(* Logix 5000 project; controller PLC_MCC1300_75F1 vendor 1 type 14 code 166 rev 32.11; software revision 32.04; part 74 of 83 *)
(* tags used below, declared in another part *)
   AUX_tConvoyCap_ZC_NULL : UDT_ConvoyCap_ZC;
   CONST_rgdDestMask : DINT[32];   // Destination Mask
   CONST_tAux : AUX_COSTANTS;
   CONST_tPlant : UDT_PLANT_CONSTANTS;
   GP_PosWindow : GP_PosWindow;
   GP_TrackingAddCap : GP_TrackingAddCap;
   M302SpeedUp : MAC_SpeedUp;
   M303_dHalfWidthDifference : DINT;
   M307ASpeedUp : MAC_SpeedUp;
   M30xTrimDeck : MAC_TrimmingDeck[5];
   M30xTrimDeck_DATA : UDT_ConvoyCap_ZC[5];
   M30xTrimDeck_HMR : MAC_TrimmingDeck_HMR[5];
   M30xTrimDeck_HMW : MAC_TrimmingDeck_HMW[5];
   M30xTrimWheel : MAC_TrimmingWheels[5];
   M310Popup : MAC_Popup_ZC[2];
   M315Popup : MAC_Popup_ZC[2];
   M350Popup : MAC_Popup_ZC;
   O : INT[128];
   Sbr_IN_dCapIndex : DINT;
   Sbr_IN_DestinationCullet : DINT;
   Sbr_IN_dIndexHead : DINT;
   Sbr_IN_ReentryPosition : DINT;
   Sbr_IN_ReentryPosition_max : DINT;
   Sbr_IN_ReentryPosition_min : DINT;
   Sbr_INO_DestinationLite : DINT;
   Sbr_INO_tConvoy_SL : UDT_Convoy_SL;
   Sbr_INO_tConvoyCap_ZC : UDT_ConvoyCap_ZC;
   Sbr_INO_xALLForDestination : BOOL;
   Sbr_INO_xAllLiteToCullet : BOOL;
   Sbr_INO_xAtLeastOneForDestination : BOOL;
   Sbr_INO_xAtLeastOneToCullet : BOOL;
   Sbr_OUT_dTotalCaps : DINT;
   Sbr_OUT_rgdConvoyGaps : DINT[4];
   Sbr_OUT_rgdConvoyLengths : DINT[4];
   TMP_d : DINT;
   TMP_dCap : DINT;
   TMP_dConvoySearchMax : DINT;
   TMP_dIndC : DINT;
   TMP_dIndex : DINT;
   TMP_dLite : DINT;
   TMP_dManualTargetPos : DINT;
   TMP_dMaxCap : DINT;
   TMP_dMaxLite : DINT;
   TMP_dNextCap : DINT;
   TMP_dPointer : DINT;
   TMP_dWander : DINT;
   TMP_rgdIndexC : DINT[4];
   TMP_rgdPnt : DINT[5];
   TMP_x : BOOL;
   TMP_xDebugOFF : BOOL;
   TMP_xDebugON : BOOL;
   xAlwaysOFF : BOOL;
   xAlwaysON : BOOL;
   Z200_SnapDataEth : UDT_ConvoyCap_ZC[2];
   Z300_BufferPlate : UDT_LINE_BUFFER_PLATE;
   Z300_Conveyor_Conf : UDT_Conveyor_Config[29];
   Z300_dEndTrackingPosition : DINT;
   Z300_LineTracking : UDT_LINE_TRACKING;
   Z301 : MAC_Zone_ML;
   Z401_HMI_rgtPlateScada : HMI_LiteData[5,2,7];
   Z401_HMI_rgtPlateScada_Internal : HMI_LiteData[5,2,7];
   Z402_HMI_rgtPlateScada : HMI_LiteData[5,2,7];
   Z402_HMI_rgtPlateScada_Internal : HMI_LiteData[5,2,7];
   Z900_HMI_rgtPlateScada : HMI_LiteData[5,2,7];
   Z900_HMI_rgtPlateScada_Internal : HMI_LiteData[5,2,7];
(* MainProgram, continued *)

ROUTINE Machines_Config   (* structured text *)
   //// MACHINES CONFIGURATION ////
   
   //M302 Speed-Up
   M302SpeedUp.AUX_dConveyorLength_cmm := 0;
   FOR TMP_dIndex := 0 TO 9 DO
   	M302SpeedUp.AUX_dConveyorLength_cmm := M302SpeedUp.AUX_dConveyorLength_cmm + Z300_Conveyor_Conf[TMP_dIndex].dLengthConveyor_cmm;
   END_FOR;
   
   //M302 Trim Deck
   M30xTrimDeck[0].CONF_dAutoSpeed_mm_min := 1000; //1680 //1000 (/60)
   M30xTrimDeck[0].CONF_dManualSpeed_mm_min := 300; //500 //900 //300 (/60)
   M30xTrimDeck[0].CONF_dConveyorLength_cmm := Z300_LineTracking.rgtTrkConv[2].dLengthConveyor + Z300_LineTracking.rgtTrkConv[3].dLengthConveyor + Z300_LineTracking.rgtTrkConv[4].dLengthConveyor + Z300_LineTracking.rgtTrkConv[5].dLengthConveyor + Z300_LineTracking.rgtTrkConv[6].dLengthConveyor;
   M30xTrimDeck[0].CONF_dStartPositionFrame := Z300_LineTracking.rgtTrkConv[2].dStartPosition_cmm;
   M30xTrimDeck[0].CONF_dStopPositionFrame_cmm := Z300_LineTracking.rgtTrkConv[6].dEndPosition_cmm;
   M30xTrimDeck[0].CONF_dTrimDeckPreset[0] := 2055; //mm
   M30xTrimDeck[0].CONF_dTrimDeckPreset[1] := 2055; //mm
   M30xTrimDeck[0].CONF_dTrimDeckCleanPos_cmm[0] := 205500;
   M30xTrimDeck[0].CONF_dTrimDeckCleanPos_cmm[1] := 205500;
   M30xTrimDeck[0].CONF_dMaxTimeToReachPosition_ms := 600;
   M30xTrimDeck[0].CONF_dTolerance_cmm := 200;
   M30xTrimDeck[0].CONF_dTrimDeckTargetWindow_cmm[0] := 200;
   M30xTrimDeck[0].CONF_dTrimDeckTargetWindow_cmm[1] := 200;
   M30xTrimDeck[0].CONF_rAcceleration_m_s2[0] := 0.06;
   M30xTrimDeck[0].CONF_rDeceleration_m_s2[0] := 0.06;
   M30xTrimDeck[0].CONF_rAcceleration_m_s2[1] := 0.06;
   M30xTrimDeck[0].CONF_rDeceleration_m_s2[1] := 0.06;
   M30xTrimDeck[0].tmOF_DriveEnable[0].PRE := 30000;
   M30xTrimDeck[0].tmOF_DriveEnable[1].PRE := 30000;
   M30xTrimDeck[0].tmON_FeedbackTimeOut[0].PRE := 5000;
   M30xTrimDeck[0].tmON_FeedbackTimeOut[1].PRE := 5000;
   M30xTrimDeck[0].tmON_FeedbackDriveReady[0].PRE := 1000;
   M30xTrimDeck[0].tmON_FeedbackDriveReady[1].PRE := 1000;
   
   //M303 Trim Deck
   M30xTrimDeck[1].CONF_dAutoSpeed_mm_min := 1000; //1680 //1000 (/60)
   M30xTrimDeck[1].CONF_dManualSpeed_mm_min := 300; //500 //900 //300 (/60)
   M30xTrimDeck[1].CONF_dConveyorLength_cmm := Z300_LineTracking.rgtTrkConv[7].dLengthConveyor + Z300_LineTracking.rgtTrkConv[8].dLengthConveyor;
   M30xTrimDeck[1].CONF_dStartPositionFrame := Z300_LineTracking.rgtTrkConv[7].dStartPosition_cmm;
   M30xTrimDeck[1].CONF_dStopPositionFrame_cmm := Z300_LineTracking.rgtTrkConv[8].dEndPosition_cmm;
   M30xTrimDeck[1].CONF_dTrimDeckPreset[0] := 2055; //mm
   M30xTrimDeck[1].CONF_dTrimDeckPreset[1] := 2055; //mm
   M30xTrimDeck[1].CONF_dTrimDeckCleanPos_cmm[0] := 205500;
   M30xTrimDeck[1].CONF_dTrimDeckCleanPos_cmm[1] := 205500;
   M30xTrimDeck[1].CONF_dMaxTimeToReachPosition_ms := 600;
   M30xTrimDeck[1].CONF_dTolerance_cmm := 200;
   M30xTrimDeck[1].CONF_dTrimDeckTargetWindow_cmm[0] := 200;
   M30xTrimDeck[1].CONF_dTrimDeckTargetWindow_cmm[1] := 200;
   M30xTrimDeck[1].CONF_rAcceleration_m_s2[0] := 0.06;
   M30xTrimDeck[1].CONF_rDeceleration_m_s2[0] := 0.06;
   M30xTrimDeck[1].CONF_rAcceleration_m_s2[1] := 0.06;
   M30xTrimDeck[1].CONF_rDeceleration_m_s2[1] := 0.06;
   M30xTrimDeck[1].tmOF_DriveEnable[0].PRE := 30000;
   M30xTrimDeck[1].tmOF_DriveEnable[1].PRE := 30000;
   M30xTrimDeck[1].tmON_FeedbackTimeOut[0].PRE := 5000;
   M30xTrimDeck[1].tmON_FeedbackTimeOut[1].PRE := 5000;
   M30xTrimDeck[1].tmON_FeedbackDriveReady[0].PRE := 1000;
   M30xTrimDeck[1].tmON_FeedbackDriveReady[1].PRE := 1000;
   
   //M304 Trim Deck
   M30xTrimDeck[2].CONF_dAutoSpeed_mm_min := 1000; //1680 //1000 (/60)
   M30xTrimDeck[2].CONF_dManualSpeed_mm_min := 300; //500 //900 //300 (/60)
   M30xTrimDeck[2].CONF_dConveyorLength_cmm := Z300_LineTracking.rgtTrkConv[9].dLengthConveyor;
   M30xTrimDeck[2].CONF_dStartPositionFrame := Z300_LineTracking.rgtTrkConv[9].dStartPosition_cmm;
   M30xTrimDeck[2].CONF_dStopPositionFrame_cmm := Z300_LineTracking.rgtTrkConv[9].dEndPosition_cmm;
   M30xTrimDeck[2].CONF_dTrimDeckPreset[0] := 2055; //mm
   M30xTrimDeck[2].CONF_dTrimDeckPreset[1] := 2055; //mm
   M30xTrimDeck[2].CONF_dTrimDeckCleanPos_cmm[0] := 205500;
   M30xTrimDeck[2].CONF_dTrimDeckCleanPos_cmm[1] := 205500;
   M30xTrimDeck[2].CONF_dMaxTimeToReachPosition_ms := 600;
   M30xTrimDeck[2].CONF_dTolerance_cmm := 200;
   M30xTrimDeck[2].CONF_dTrimDeckTargetWindow_cmm[0] := 200;
   M30xTrimDeck[2].CONF_dTrimDeckTargetWindow_cmm[1] := 200;
   M30xTrimDeck[2].CONF_rAcceleration_m_s2[0] := 0.06;
   M30xTrimDeck[2].CONF_rDeceleration_m_s2[0] := 0.06;
   M30xTrimDeck[2].CONF_rAcceleration_m_s2[1] := 0.06;
   M30xTrimDeck[2].CONF_rDeceleration_m_s2[1] := 0.06;
   M30xTrimDeck[2].tmOF_DriveEnable[0].PRE := 30000;
   M30xTrimDeck[2].tmOF_DriveEnable[1].PRE := 30000;
   M30xTrimDeck[2].tmON_FeedbackTimeOut[0].PRE := 5000;
   M30xTrimDeck[2].tmON_FeedbackTimeOut[1].PRE := 5000;
   M30xTrimDeck[2].tmON_FeedbackDriveReady[0].PRE := 1000;
   M30xTrimDeck[2].tmON_FeedbackDriveReady[1].PRE := 1000;
   
   //M305 Trim Deck
   M30xTrimDeck[3].CONF_dAutoSpeed_mm_min := 1000; //1680 //1000 (/60)
   M30xTrimDeck[3].CONF_dManualSpeed_mm_min := 300; //500 //900 //300 (/60)
   M30xTrimDeck[3].CONF_dConveyorLength_cmm := Z300_LineTracking.rgtTrkConv[10].dLengthConveyor;
   M30xTrimDeck[3].CONF_dStartPositionFrame := Z300_LineTracking.rgtTrkConv[10].dStartPosition_cmm;
   M30xTrimDeck[3].CONF_dStopPositionFrame_cmm := Z300_LineTracking.rgtTrkConv[10].dEndPosition_cmm;
   M30xTrimDeck[3].CONF_dTrimDeckPreset[0] := 2055; //mm
   M30xTrimDeck[3].CONF_dTrimDeckPreset[1] := 2055; //mm
   M30xTrimDeck[3].CONF_dTrimDeckCleanPos_cmm[0] := 205500;
   M30xTrimDeck[3].CONF_dTrimDeckCleanPos_cmm[1] := 205500;
   M30xTrimDeck[3].CONF_dMaxTimeToReachPosition_ms := 600;
   M30xTrimDeck[3].CONF_dTolerance_cmm := 200;
   M30xTrimDeck[3].CONF_dTrimDeckTargetWindow_cmm[0] := 200;
   M30xTrimDeck[3].CONF_dTrimDeckTargetWindow_cmm[1] := 200;
   M30xTrimDeck[3].CONF_rAcceleration_m_s2[0] := 0.06;
   M30xTrimDeck[3].CONF_rDeceleration_m_s2[0] := 0.06;
   M30xTrimDeck[3].CONF_rAcceleration_m_s2[1] := 0.06;
   M30xTrimDeck[3].CONF_rDeceleration_m_s2[1] := 0.06;
   M30xTrimDeck[3].tmOF_DriveEnable[0].PRE := 30000;
   M30xTrimDeck[3].tmOF_DriveEnable[1].PRE := 30000;
   M30xTrimDeck[3].tmON_FeedbackTimeOut[0].PRE := 5000;
   M30xTrimDeck[3].tmON_FeedbackTimeOut[1].PRE := 5000;
   M30xTrimDeck[3].tmON_FeedbackDriveReady[0].PRE := 1000;
   M30xTrimDeck[3].tmON_FeedbackDriveReady[1].PRE := 1000;
   
   //M306 Trim Deck
   M30xTrimDeck[4].CONF_dAutoSpeed_mm_min := 1000; //1680 //1000 (/60)
   M30xTrimDeck[4].CONF_dManualSpeed_mm_min := 300; //500 //900 //300 (/60)
   M30xTrimDeck[4].CONF_dConveyorLength_cmm := Z300_LineTracking.rgtTrkConv[11].dLengthConveyor;
   M30xTrimDeck[4].CONF_dStartPositionFrame := Z300_LineTracking.rgtTrkConv[11].dStartPosition_cmm;
   M30xTrimDeck[4].CONF_dStopPositionFrame_cmm := Z300_LineTracking.rgtTrkConv[11].dEndPosition_cmm;
   M30xTrimDeck[4].CONF_dTrimDeckPreset[0] := 2055; //mm
   M30xTrimDeck[4].CONF_dTrimDeckPreset[1] := 2055; //mm
   M30xTrimDeck[4].CONF_dTrimDeckCleanPos_cmm[0] := 205500;
   M30xTrimDeck[4].CONF_dTrimDeckCleanPos_cmm[1] := 205500;
   M30xTrimDeck[4].CONF_dMaxTimeToReachPosition_ms := 600;
   M30xTrimDeck[4].CONF_dTolerance_cmm := 200;
   M30xTrimDeck[4].CONF_dTrimDeckTargetWindow_cmm[0] := 200;
   M30xTrimDeck[4].CONF_dTrimDeckTargetWindow_cmm[1] := 200;
   M30xTrimDeck[4].CONF_rAcceleration_m_s2[0] := 0.06;
   M30xTrimDeck[4].CONF_rDeceleration_m_s2[0] := 0.06;
   M30xTrimDeck[4].CONF_rAcceleration_m_s2[1] := 0.06;
   M30xTrimDeck[4].CONF_rDeceleration_m_s2[1] := 0.06;
   M30xTrimDeck[4].tmOF_DriveEnable[0].PRE := 30000;
   M30xTrimDeck[4].tmOF_DriveEnable[1].PRE := 30000;
   M30xTrimDeck[4].tmON_FeedbackTimeOut[0].PRE := 5000;
   M30xTrimDeck[4].tmON_FeedbackTimeOut[1].PRE := 5000;
   M30xTrimDeck[4].tmON_FeedbackDriveReady[0].PRE := 1000;
   M30xTrimDeck[4].tmON_FeedbackDriveReady[1].PRE := 1000;
   
   //M302 Trim Wheels
   M30xTrimWheel[0].CONF_dAutoSpeed_mm_min[0] := 1000;
   M30xTrimWheel[0].CONF_dAutoSpeed_mm_min[1] := 1000;
   M30xTrimWheel[0].CONF_dManualSpeed_mm_min[0] := 200;
   M30xTrimWheel[0].CONF_dManualSpeed_mm_min[1] := 200;
   M30xTrimWheel[0].CONF_dAutoSpeed_mm_min[1] := 1000;
   M30xTrimWheel[0].CONF_dMaxTimeToReachPosition_ms[0] := 600;
   M30xTrimWheel[0].CONF_dMaxTimeToReachPosition_ms[1] := 600;
   M30xTrimWheel[0].CONF_dTolerance_cmm[0] := 200;
   M30xTrimWheel[0].CONF_dTolerance_cmm[1] := 200;
   M30xTrimWheel[0].CONF_dTrimWheelTargetWindow_cmm[0] := 200;
   M30xTrimWheel[0].CONF_dTrimWheelTargetWindow_cmm[1] := 200;
   M30xTrimWheel[0].CONF_dTrimWheelMinPos_cmm[0] := 115000;
   M30xTrimWheel[0].CONF_dTrimWheelMinPos_cmm[1] := 115000;
   M30xTrimWheel[0].CONF_dTrimWheelMaxPos_cmm[0] := 262000;
   M30xTrimWheel[0].CONF_dTrimWheelMaxPos_cmm[1] := 256000;
   M30xTrimWheel[0].CONF_dTrimWheelMinRange_cmm[0] := 115000;
   M30xTrimWheel[0].CONF_dTrimWheelMinRange_cmm[1] := 115000;
   M30xTrimWheel[0].CONF_dTrimWheelMaxRange_cmm[0] := 262000;
   M30xTrimWheel[0].CONF_dTrimWheelMaxRange_cmm[1] := 256000;
   M30xTrimWheel[0].CONF_dTrimWheelCodeOpt := 1;
   M30xTrimWheel[0].CONF_dConveyorLength_cmm := Z300_LineTracking.rgtTrkConv[2].dLengthConveyor;
   M30xTrimWheel[0].CONF_dMaxLengthWorkable_cmm := 680000;
   M30xTrimWheel[0].CONF_dPositionWheel_cmm := Z300_LineTracking.rgtTrkConv[2].dEndPosition_cmm;
   M30xTrimWheel[0].CONF_dTrimWheelArmPos_cmm[0] := Z300_LineTracking.rgtTrkConv[2].dEndPosition_cmm;
   M30xTrimWheel[0].CONF_dTrimWheelArmPos_cmm[1] := Z300_LineTracking.rgtTrkConv[2].dEndPosition_cmm;
   M30xTrimWheel[0].CONF_rAcceleration_m_s2[0] := 1.0;
   M30xTrimWheel[0].CONF_rAcceleration_m_s2[1] := 1.0;
   M30xTrimWheel[0].CONF_rDeceleration_m_s2[0] := 1.0;
   M30xTrimWheel[0].CONF_rDeceleration_m_s2[1] := 1.0;
   M30xTrimWheel[0].CONF_dTrimWheelPresetZero_cmm[0] := 2055; //(1905+150) //mm
   M30xTrimWheel[0].CONF_dTrimWheelPresetZero_cmm[1] := 2055; //(1905+150) //mm
   M30xTrimWheel[0].tmOF_DriveEnable[0].PRE := 30000;
   M30xTrimWheel[0].tmOF_DriveEnable[1].PRE := 30000;
   M30xTrimWheel[0].tmON_FeedbackTimeOut[0].PRE := 3500;
   M30xTrimWheel[0].tmON_FeedbackTimeOut[1].PRE := 3500;
   M30xTrimWheel[0].tmON_FeedbackDriveReady[0].PRE := 1000;
   M30xTrimWheel[0].tmON_FeedbackDriveReady[1].PRE := 1000;
   
   //M303 Trim Wheels
   M30xTrimWheel[1].CONF_dAutoSpeed_mm_min[0] := 1000;
   M30xTrimWheel[1].CONF_dAutoSpeed_mm_min[1] := 1000;
   M30xTrimWheel[1].CONF_dManualSpeed_mm_min[0] := 200;
   M30xTrimWheel[1].CONF_dManualSpeed_mm_min[1] := 200;
   M30xTrimWheel[1].CONF_dAutoSpeed_mm_min[1] := 1000;
   M30xTrimWheel[1].CONF_dMaxTimeToReachPosition_ms[0] := 600;
   M30xTrimWheel[1].CONF_dMaxTimeToReachPosition_ms[1] := 600;
   M30xTrimWheel[1].CONF_dTolerance_cmm[0] := 200;
   M30xTrimWheel[1].CONF_dTolerance_cmm[1] := 200;
   M30xTrimWheel[1].CONF_dTrimWheelTargetWindow_cmm[0] := 200;
   M30xTrimWheel[1].CONF_dTrimWheelTargetWindow_cmm[1] := 200;
   M30xTrimWheel[1].CONF_dTrimWheelMinPos_cmm[0] := -15000;
   M30xTrimWheel[1].CONF_dTrimWheelMinPos_cmm[1] := -15000;
   M30xTrimWheel[1].CONF_dTrimWheelMaxPos_cmm[0] := 42000;
   M30xTrimWheel[1].CONF_dTrimWheelMaxPos_cmm[1] := 42000;
   M30xTrimWheel[1].CONF_dTrimWheelMinRange_cmm[0] := -15000;
   M30xTrimWheel[1].CONF_dTrimWheelMinRange_cmm[1] := -15000;
   M30xTrimWheel[1].CONF_dTrimWheelMaxRange_cmm[0] := 42000;
   M30xTrimWheel[1].CONF_dTrimWheelMaxRange_cmm[1] := 42000;
   M30xTrimWheel[1].CONF_dTrimWheelCodeOpt := 2;
   M30xTrimWheel[1].CONF_dConveyorLength_cmm := Z300_LineTracking.rgtTrkConv[7].dLengthConveyor + Z300_LineTracking.rgtTrkConv[8].dLengthConveyor;
   M30xTrimWheel[1].CONF_dMaxLengthWorkable_cmm := 610000;
   M30xTrimWheel[1].CONF_dPositionWheel_cmm := Z300_LineTracking.rgtTrkConv[8].dEndPosition_cmm - 8000;
   M30xTrimWheel[1].CONF_dTrimWheelArmPos_cmm[0] := Z300_LineTracking.rgtTrkConv[8].dEndPosition_cmm - 8000;
   M30xTrimWheel[1].CONF_dTrimWheelArmPos_cmm[1] := Z300_LineTracking.rgtTrkConv[8].dEndPosition_cmm - 8000;
   M30xTrimWheel[1].CONF_rAcceleration_m_s2[0] := 1.0;
   M30xTrimWheel[1].CONF_rAcceleration_m_s2[1] := 1.0;
   M30xTrimWheel[1].CONF_rDeceleration_m_s2[0] := 1.0;
   M30xTrimWheel[1].CONF_rDeceleration_m_s2[1] := 1.0;
   M30xTrimWheel[1].CONF_dTrimWheelPresetZero_cmm[0] := 2055; //(1905+150) //mm
   M30xTrimWheel[1].CONF_dTrimWheelPresetZero_cmm[1] := 2055; //(1905+150) //mm
   M30xTrimWheel[1].tmOF_DriveEnable[0].PRE := 30000;
   M30xTrimWheel[1].tmOF_DriveEnable[1].PRE := 30000;
   M30xTrimWheel[1].tmON_FeedbackTimeOut[0].PRE := 3500;
   M30xTrimWheel[1].tmON_FeedbackTimeOut[1].PRE := 3500;
   M30xTrimWheel[1].tmON_FeedbackDriveReady[0].PRE := 1000;
   M30xTrimWheel[1].tmON_FeedbackDriveReady[1].PRE := 1000;
   ////These trimming wheels work on tail position
   //M303xTrimWheel[1].ST_xTailBreakOpSide := 1;
   //M303xTrimWheel[1].ST_xTailBreakOppOpSide := 1;
   
   //M304 Trim Wheels
   M30xTrimWheel[2].CONF_dAutoSpeed_mm_min[0] := 1000;
   M30xTrimWheel[2].CONF_dAutoSpeed_mm_min[1] := 1000;
   M30xTrimWheel[2].CONF_dManualSpeed_mm_min[0] := 200;
   M30xTrimWheel[2].CONF_dManualSpeed_mm_min[1] := 200;
   M30xTrimWheel[2].CONF_dAutoSpeed_mm_min[1] := 1000;
   M30xTrimWheel[2].CONF_dMaxTimeToReachPosition_ms[0] := 600;
   M30xTrimWheel[2].CONF_dMaxTimeToReachPosition_ms[1] := 600;
   M30xTrimWheel[2].CONF_dTolerance_cmm[0] := 200;
   M30xTrimWheel[2].CONF_dTolerance_cmm[1] := 200;
   M30xTrimWheel[2].CONF_dTrimWheelTargetWindow_cmm[0] := 200;
   M30xTrimWheel[2].CONF_dTrimWheelTargetWindow_cmm[1] := 200;
   M30xTrimWheel[2].CONF_dTrimWheelMinPos_cmm[0] := -15000;
   M30xTrimWheel[2].CONF_dTrimWheelMinPos_cmm[1] := -15000;
   M30xTrimWheel[2].CONF_dTrimWheelMaxPos_cmm[0] := 42000;
   M30xTrimWheel[2].CONF_dTrimWheelMaxPos_cmm[1] := 42000;
   M30xTrimWheel[2].CONF_dTrimWheelMinRange_cmm[0] := -15000;
   M30xTrimWheel[2].CONF_dTrimWheelMinRange_cmm[1] := -15000;
   M30xTrimWheel[2].CONF_dTrimWheelMaxRange_cmm[0] := 42000;
   M30xTrimWheel[2].CONF_dTrimWheelMaxRange_cmm[1] := 42000;
   M30xTrimWheel[2].CONF_dTrimWheelCodeOpt := 3;
   M30xTrimWheel[2].CONF_dConveyorLength_cmm := Z300_LineTracking.rgtTrkConv[9].dLengthConveyor;
   M30xTrimWheel[2].CONF_dMaxLengthWorkable_cmm := 680000;
   M30xTrimWheel[2].CONF_dPositionWheel_cmm := Z300_LineTracking.rgtTrkConv[9].dEndPosition_cmm - 8000;
   M30xTrimWheel[2].CONF_dTrimWheelArmPos_cmm[0] := Z300_LineTracking.rgtTrkConv[9].dEndPosition_cmm - 8000;
   M30xTrimWheel[2].CONF_dTrimWheelArmPos_cmm[1] := Z300_LineTracking.rgtTrkConv[9].dEndPosition_cmm - 8000;
   M30xTrimWheel[2].CONF_rAcceleration_m_s2[0] := 1.0;
   M30xTrimWheel[2].CONF_rAcceleration_m_s2[1] := 1.0;
   M30xTrimWheel[2].CONF_rDeceleration_m_s2[0] := 1.0;
   M30xTrimWheel[2].CONF_rDeceleration_m_s2[1] := 1.0;
   M30xTrimWheel[2].CONF_dTrimWheelPresetZero_cmm[0] := 2055; //(1905+150) //mm
   M30xTrimWheel[2].CONF_dTrimWheelPresetZero_cmm[1] := 2055; //(1905+150) //mm
   M30xTrimWheel[2].tmOF_DriveEnable[0].PRE := 30000;
   M30xTrimWheel[2].tmOF_DriveEnable[1].PRE := 30000;
   M30xTrimWheel[2].tmON_FeedbackTimeOut[0].PRE := 3500;
   M30xTrimWheel[2].tmON_FeedbackTimeOut[1].PRE := 3500;
   M30xTrimWheel[2].tmON_FeedbackDriveReady[0].PRE := 1000;
   M30xTrimWheel[2].tmON_FeedbackDriveReady[1].PRE := 1000;
   
   //M305 Trim Wheels
   M30xTrimWheel[3].CONF_dAutoSpeed_mm_min[0] := 1000;
   M30xTrimWheel[3].CONF_dAutoSpeed_mm_min[1] := 1000;
   M30xTrimWheel[3].CONF_dManualSpeed_mm_min[0] := 200;
   M30xTrimWheel[3].CONF_dManualSpeed_mm_min[1] := 200;
   M30xTrimWheel[3].CONF_dAutoSpeed_mm_min[1] := 1000;
   M30xTrimWheel[3].CONF_dMaxTimeToReachPosition_ms[0] := 600;
   M30xTrimWheel[3].CONF_dMaxTimeToReachPosition_ms[1] := 600;
   M30xTrimWheel[3].CONF_dTolerance_cmm[0] := 200;
   M30xTrimWheel[3].CONF_dTolerance_cmm[1] := 200;
   M30xTrimWheel[3].CONF_dTrimWheelTargetWindow_cmm[0] := 200;
   M30xTrimWheel[3].CONF_dTrimWheelTargetWindow_cmm[1] := 200;
   M30xTrimWheel[3].CONF_dTrimWheelMinPos_cmm[0] := -15000;
   M30xTrimWheel[3].CONF_dTrimWheelMinPos_cmm[1] := -15000;
   M30xTrimWheel[3].CONF_dTrimWheelMaxPos_cmm[0] := 42000;
   M30xTrimWheel[3].CONF_dTrimWheelMaxPos_cmm[1] := 42000;
   M30xTrimWheel[3].CONF_dTrimWheelMinRange_cmm[0] := -15000;
   M30xTrimWheel[3].CONF_dTrimWheelMinRange_cmm[1] := -15000;
   M30xTrimWheel[3].CONF_dTrimWheelMaxRange_cmm[0] := 42000;
   M30xTrimWheel[3].CONF_dTrimWheelMaxRange_cmm[1] := 42000;
   M30xTrimWheel[3].CONF_dTrimWheelCodeOpt := 4;
   M30xTrimWheel[3].CONF_dConveyorLength_cmm := Z300_LineTracking.rgtTrkConv[10].dLengthConveyor;
   M30xTrimWheel[3].CONF_dMaxLengthWorkable_cmm := 610000;
   M30xTrimWheel[3].CONF_dPositionWheel_cmm := Z300_LineTracking.rgtTrkConv[10].dEndPosition_cmm - 8000;
   M30xTrimWheel[3].CONF_dTrimWheelArmPos_cmm[0] := Z300_LineTracking.rgtTrkConv[10].dEndPosition_cmm - 8000;
   M30xTrimWheel[3].CONF_dTrimWheelArmPos_cmm[1] := Z300_LineTracking.rgtTrkConv[10].dEndPosition_cmm - 8000;
   M30xTrimWheel[3].CONF_rAcceleration_m_s2[0] := 1.0;
   M30xTrimWheel[3].CONF_rAcceleration_m_s2[1] := 1.0;
   M30xTrimWheel[3].CONF_rDeceleration_m_s2[0] := 1.0;
   M30xTrimWheel[3].CONF_rDeceleration_m_s2[1] := 1.0;
   M30xTrimWheel[3].CONF_dTrimWheelPresetZero_cmm[0] := 2055; //(1905+150) //mm
   M30xTrimWheel[3].CONF_dTrimWheelPresetZero_cmm[1] := 2055; //(1905+150) //mm
   M30xTrimWheel[3].tmOF_DriveEnable[0].PRE := 30000;
   M30xTrimWheel[3].tmOF_DriveEnable[1].PRE := 30000;
   M30xTrimWheel[3].tmON_FeedbackTimeOut[0].PRE := 3500;
   M30xTrimWheel[3].tmON_FeedbackTimeOut[1].PRE := 3500;
   M30xTrimWheel[3].tmON_FeedbackDriveReady[0].PRE := 1000;
   M30xTrimWheel[3].tmON_FeedbackDriveReady[1].PRE := 1000;
   
   //M306 Trim Wheels
   M30xTrimWheel[4].CONF_dAutoSpeed_mm_min[0] := 1000;
   M30xTrimWheel[4].CONF_dAutoSpeed_mm_min[1] := 1000;
   M30xTrimWheel[4].CONF_dManualSpeed_mm_min[0] := 200;
   M30xTrimWheel[4].CONF_dManualSpeed_mm_min[1] := 200;
   M30xTrimWheel[4].CONF_dAutoSpeed_mm_min[1] := 1000;
   M30xTrimWheel[4].CONF_dMaxTimeToReachPosition_ms[0] := 600;
   M30xTrimWheel[4].CONF_dMaxTimeToReachPosition_ms[1] := 600;
   M30xTrimWheel[4].CONF_dTolerance_cmm[0] := 200;
   M30xTrimWheel[4].CONF_dTolerance_cmm[1] := 200;
   M30xTrimWheel[4].CONF_dTrimWheelTargetWindow_cmm[0] := 200;
   M30xTrimWheel[4].CONF_dTrimWheelTargetWindow_cmm[1] := 200;
   M30xTrimWheel[4].CONF_dTrimWheelMinPos_cmm[0] := -15000;
   M30xTrimWheel[4].CONF_dTrimWheelMinPos_cmm[1] := -15000;
   M30xTrimWheel[4].CONF_dTrimWheelMaxPos_cmm[0] := 42000;
   M30xTrimWheel[4].CONF_dTrimWheelMaxPos_cmm[1] := 42000;
   M30xTrimWheel[4].CONF_dTrimWheelMinRange_cmm[0] := -15000;
   M30xTrimWheel[4].CONF_dTrimWheelMinRange_cmm[1] := -15000;
   M30xTrimWheel[4].CONF_dTrimWheelMaxRange_cmm[0] := 42000;
   M30xTrimWheel[4].CONF_dTrimWheelMaxRange_cmm[1] := 42000;
   M30xTrimWheel[4].CONF_dTrimWheelCodeOpt := 4;
   M30xTrimWheel[4].CONF_dConveyorLength_cmm := Z300_LineTracking.rgtTrkConv[11].dLengthConveyor;
   M30xTrimWheel[4].CONF_dMaxLengthWorkable_cmm := 610000;
   M30xTrimWheel[4].CONF_dPositionWheel_cmm := Z300_LineTracking.rgtTrkConv[11].dEndPosition_cmm - 8000;
   M30xTrimWheel[4].CONF_dTrimWheelArmPos_cmm[0] := Z300_LineTracking.rgtTrkConv[11].dEndPosition_cmm - 8000;
   M30xTrimWheel[4].CONF_dTrimWheelArmPos_cmm[1] := Z300_LineTracking.rgtTrkConv[11].dEndPosition_cmm - 8000;
   M30xTrimWheel[4].CONF_rAcceleration_m_s2[0] := 1.0;
   M30xTrimWheel[4].CONF_rAcceleration_m_s2[1] := 1.0;
   M30xTrimWheel[4].CONF_rDeceleration_m_s2[0] := 1.0;
   M30xTrimWheel[4].CONF_rDeceleration_m_s2[1] := 1.0;
   M30xTrimWheel[4].CONF_dTrimWheelPresetZero_cmm[0] := 2055; //(1905+150) //mm
   M30xTrimWheel[4].CONF_dTrimWheelPresetZero_cmm[1] := 2055; //(1905+150) //mm
   M30xTrimWheel[4].tmOF_DriveEnable[0].PRE := 30000;
   M30xTrimWheel[4].tmOF_DriveEnable[1].PRE := 30000;
   M30xTrimWheel[4].tmON_FeedbackTimeOut[0].PRE := 3500;
   M30xTrimWheel[4].tmON_FeedbackTimeOut[1].PRE := 3500;
   M30xTrimWheel[4].tmON_FeedbackDriveReady[0].PRE := 1000;
   M30xTrimWheel[4].tmON_FeedbackDriveReady[1].PRE := 1000;
   
   
   //M307A Speed-Up
   M307ASpeedUp.AUX_dConveyorLength_cmm := 0;
   FOR TMP_dIndex := 8 TO 10 DO
   	M307ASpeedUp.AUX_dConveyorLength_cmm := M307ASpeedUp.AUX_dConveyorLength_cmm + Z300_Conveyor_Conf[TMP_dIndex].dLengthConveyor_cmm;
   END_FOR;
   
   //M350Popup
   M350Popup.AUX_dPosTimeout := M350Popup.AUX_dEndPosition_cmm + 400000;
   
   //M310Popup
   M310Popup[0].AUX_dPosTimeout := M310Popup[0].AUX_dEndPosition_cmm + 600000;
   M310Popup[1].AUX_dPosTimeout := M310Popup[1].AUX_dEndPosition_cmm + 400000;
   
   //M315Popup
   M315Popup[0].AUX_dPosTimeout := M315Popup[0].AUX_dEndPosition_cmm + 800000;
   M315Popup[1].AUX_dPosTimeout := M315Popup[1].AUX_dEndPosition_cmm + 400000;
   
END_ROUTINE

ROUTINE MainRoutine   (* ladder *)
   0: [OTU(xAlwaysOFF) ,OTU(TMP_xDebugOFF) ];
   1: XIO(xAlwaysOFF)[OTL(xAlwaysON) ,OTL(TMP_xDebugON) ];
   2: XIC(TMP_xDebugOFF)JSR(_812_HOST_MOVE,1,500)JSR(_814_HOST_MOVE,1,999);
   3: JSR(inputs_update,0);
   4: JSR(_2_MCP_A,0)JSR(_3_MCP_B,0);
   5: JSR(_7_MCP_F,0)JSR(_9_MCP_H,0)JSR(_10_MCP_I,0)JSR(_12_MCP_K,0);
   6: JSR(Conv_Config,0);
   7: JSR(Machines_Config,0);
   8: JSR(Conv_Mapping,0);
   9: JSR(Tracking_Logic,0);
   10: JSR(Z301_Logic,0);
   11: JSR(Conv_Main,0);
   12: JSR(ScadaPlate_Logic,0);
   13: JSR(M302SpeedUp_Logic,0);
   14: FOR(M30xTrimDeckManagement,TMP_dIndex,0,4,1);
   15: FOR(M30xTrimDeck_Logic,TMP_dIndex,0,4,1);
   16: FOR(M30xTrimWheelBrManagement,TMP_dIndex,0,4,1);
   17: FOR(M30xTrimWheelTrManagement,TMP_dIndex,0,4,1);
   18: FOR(M30xTrimWheel_Logic,TMP_dIndex,0,4,1);
   19: JSR(Hold_Down_Wheels,0);
   20: JSR(_4_VIS_INTFCE,0);
   21: JSR(M307ASpeedUp_Logic,0);
   22: JSR(M350PopupManagement,0);
   23: JSR(M350Popup_Logic,0);
   24: JSR(M310PopupManagement,0);
   25: JSR(M310Popup0_Logic,0);
   26: JSR(M310Popup1_Logic,0);
   27: JSR(M315PopupManagement,0);
   28: JSR(M315Popup0_Logic,0);
   29: JSR(M315Popup1_Logic,0);
   30: FLL(0,Z401_HMI_rgtPlateScada_Internal[0,0,0],70);
   31: FLL(0,Z402_HMI_rgtPlateScada_Internal[0,0,0],70);
   32: FLL(0,Z900_HMI_rgtPlateScada_Internal[0,0,0],70);
   33: JSR(Z401_Logic,0);
   34: JSR(M310B_Logic,0);
   35: JSR(Z311S_Logic,0);
   36: JSR(M311_Logic,0);
   37: JSR(M312_Logic,0);
   38: JSR(Z402_Logic,0);
   39: JSR(M315B_Logic,0);
   40: JSR(M315A_Logic,0);
   41: JSR(M316_Logic,0);
   42: JSR(Z316S_Logic,0);
   43: JSR(M317_Logic,0);
   44: JSR(Z900_Logic,0);
   45: JSR(M351_Logic,0);
   46: JSR(M352_Logic,0);
   47: COP(Z401_HMI_rgtPlateScada_Internal[0,0,0],Z401_HMI_rgtPlateScada[0,0,0],70);
   48: COP(Z402_HMI_rgtPlateScada_Internal[0,0,0],Z402_HMI_rgtPlateScada[0,0,0],70);
   49: COP(Z900_HMI_rgtPlateScada_Internal[0,0,0],Z900_HMI_rgtPlateScada[0,0,0],70);
   50: JSR(_811_HOST_MOVE,1,500);
   51: JSR(outputs_update,0);
END_ROUTINE

ROUTINE outputs_update   (* ladder *)
   0: COP(O[9],ETH_M2:11:O.Data,1);
   1: COP(O[16],VMCC_TD:O.Data[0],8)COP(O[24],ROCKWELL_CAPPING_SYSTEM:O.Data[0],2)COP(O[26],VMCC_M2CM01_SPEED:O.Data[0],2)COP(O[28],VMCC_M2_M2CM02_Speed:O.Data[0],2)COP(O[30],VMCC_M2_M2CM03_Speed:O.Data[0],2);
   2: COP(O[32],PANEL_KD_CS1N:O.Data[0],4)COP(O[36],PANEL_TD_CS1N:O.Data[0],4);
   3: COP(O[40],Panel_TS_CS2N:O.Data[0],4)COP(O[44],PANEL_TD_CS3N:O.Data[0],4);
   4: COP(O[48],PANEL_TD_CS4N:O.Data[0],4)COP(O[52],PANEL_TD_CS5N:O.Data[0],4);
   5: COP(O[56],PANEL_TD_CS5S:O.Data[0],4)COP(O[60],PANEL_TD_CS4S:O.Data[0],4);
   6: COP(O[64],PANEL_TD_CS3S:O.Data[0],4)COP(O[68],PANEL_TD_CS2S:O.Data[0],4);
   7: COP(O[72],BENCHBOARD:O.Data[0],4)COP(O[76],PANEL_KD_CS1S:O.Data[0],4);
   8: COP(O[80],PANEL_TD_CS1S:O.Data[0],4)COP(O[84],VMCC_M2CM4S:O.Data[0],2)COP(O[86],VMCC_M2_M2CM4N:O.Data[0],2);
   9: COP(O[104],VMCC_M2_M2CM9S:O.Data[0],2)COP(O[106],VMCC_M2_M2CM9N:O.Data[0],2)COP(O[108],VMCC_M2_M2CM10S:O.Data[0],2)COP(O[110],VMCC_M2_M2CM10N:O.Data[0],2);
   10: COP(O[112],VMCC_M2_M2CM11S:O.Data[0],2)COP(O[114],VMCC_M2_M2CM11N:O.Data[0],2)COP(O[116],VMCC_M2_M2CM12S:O.Data[0],2)COP(O[118],VMCC_M2_M2CM12N:O.Data[0],2);
   11: COP(O[120],MB:O.Data[0],8);
   12: COP(O[88],VMCC_M2_M2CM5S:O.Data[0],2)COP(O[90],VMCC_M2_M2CM5N:O.Data[0],2)COP(O[92],VMCC_M2_M2CM6S:O.Data[0],2)COP(O[94],VMCC_M2_M2CM6N:O.Data[0],2);
   13: COP(O[96],VMCC_M2_M2CM7S:O.Data[0],2)COP(O[98],VMCC_M2_M2CM7N:O.Data[0],2)COP(O[100],VMCC_M2_M2CM8S:O.Data[0],2)COP(O[102],VMCC_M2_M2CM8N:O.Data[0],2);
END_ROUTINE

ROUTINE sbrCheckConvoySLDestination   (* structured text *)
   
   SBR(Sbr_INO_tConvoy_SL,Sbr_INO_DestinationLite,Sbr_IN_DestinationCullet);
   
   SIZE(Sbr_INO_tConvoy_SL.rgtCap[0],0,TMP_dMaxCap);
   SIZE(Sbr_INO_tConvoy_SL.rgtCap[0].rgtLite[0],0,TMP_dMaxLite);
   
   Sbr_INO_xAllLiteToCullet := 1;
   Sbr_INO_xAtLeastOneForDestination := 0;
   FOR TMP_dCap := 0 TO TMP_dMaxCap - 1 DO
   	FOR TMP_dLite := 0 TO TMP_dMaxLite - 1 DO
   		IF Sbr_INO_tConvoy_SL.rgtCap[TMP_dCap].rgtLite[TMP_dLite].dID <> 0 THEN
   			IF Sbr_INO_tConvoy_SL.rgtCap[TMP_dCap].rgtLite[TMP_dLite].tDestination.rgxMain = Sbr_INO_DestinationLite THEN
   				Sbr_INO_xAtLeastOneForDestination := 1;
   			END_IF;
   			IF NOT (Sbr_INO_tConvoy_SL.rgtCap[TMP_dCap].rgtLite[TMP_dLite].tDestination.rgxMain = Sbr_IN_DestinationCullet) THEN
   				Sbr_INO_xAllLiteToCullet := 0;
   			END_IF;
   		END_IF;
   	END_FOR;
   END_FOR;
   
   RET(Sbr_INO_xAllLiteToCullet,Sbr_INO_xAtLeastOneForDestination);
END_ROUTINE

ROUTINE sbrCheckConvoyZCDestination   (* structured text *)
   
   SBR(Sbr_IN_dCapIndex,Sbr_INO_DestinationLite,Sbr_IN_DestinationCullet,Sbr_INO_xAtLeastOneForDestination,Sbr_INO_xAllLiteToCullet);
   
   FOR TMP_dLite := 0 TO Z300_BufferPlate.rgtPlate[Sbr_IN_dCapIndex].tData.rgtCap[0].dNumLites - 1 DO
   	IF Z300_BufferPlate.rgtPlate[Sbr_IN_dCapIndex].tData.rgtCap[0].rgtLite[TMP_dLite].dID <> 0 THEN
   		IF Z300_BufferPlate.rgtPlate[Sbr_IN_dCapIndex].tData.rgtCap[0].rgtLite[TMP_dLite].tDestination.rgxMain = Sbr_INO_DestinationLite THEN
   			Sbr_INO_xAtLeastOneForDestination := 1;
   		END_IF;
   		IF NOT (Z300_BufferPlate.rgtPlate[Sbr_IN_dCapIndex].tData.rgtCap[0].rgtLite[TMP_dLite].tDestination.rgxMain = Sbr_IN_DestinationCullet) THEN
   			Sbr_INO_xAllLiteToCullet := 0;
   		END_IF;
   	END_IF;
   END_FOR;
   TMP_dNextCap := Z300_BufferPlate.rgtPlate[Sbr_IN_dCapIndex].tTracking.dNextCapIndex;
   IF (Z300_BufferPlate.rgtPlate[Sbr_IN_dCapIndex].tData.dTotalCaps > 1) AND (TMP_dNextCap > 0) THEN
   	JSR(sbrCheckConvoyZCDestination,5,TMP_dNextCap,Sbr_INO_DestinationLite,Sbr_IN_DestinationCullet,Sbr_INO_xAtLeastOneForDestination,Sbr_INO_xAllLiteToCullet,Sbr_INO_xAtLeastOneForDestination,Sbr_INO_xAllLiteToCullet);
   END_IF;
   
   RET(Sbr_INO_xAtLeastOneForDestination,Sbr_INO_xAllLiteToCullet);
   
END_ROUTINE

ROUTINE sbrCheckConvoyZCDestinationFull   (* structured text *)
   
   
   SBR(Sbr_IN_dCapIndex,Sbr_INO_DestinationLite,Sbr_IN_DestinationCullet,Sbr_INO_xALLForDestination,Sbr_INO_xAtLeastOneToCullet);
   
   FOR TMP_dLite := 0 TO Z300_BufferPlate.rgtPlate[Sbr_IN_dCapIndex].tData.rgtCap[0].dNumLites - 1 DO
   	IF Z300_BufferPlate.rgtPlate[Sbr_IN_dCapIndex].tData.rgtCap[0].rgtLite[TMP_dLite].dID <> 0 THEN
   		IF NOT (Z300_BufferPlate.rgtPlate[Sbr_IN_dCapIndex].tData.rgtCap[0].rgtLite[TMP_dLite].tDestination.rgxMain = Sbr_INO_DestinationLite) THEN
   			Sbr_INO_xALLForDestination := 0;
   		END_IF;
   		IF (Z300_BufferPlate.rgtPlate[Sbr_IN_dCapIndex].tData.rgtCap[0].rgtLite[TMP_dLite].tDestination.rgxMain = Sbr_IN_DestinationCullet) THEN
   			Sbr_INO_xAtLeastOneToCullet := 1;
   		END_IF;
   	END_IF;
   END_FOR;
   TMP_dNextCap := Z300_BufferPlate.rgtPlate[Sbr_IN_dCapIndex].tTracking.dNextCapIndex;
   IF (Z300_BufferPlate.rgtPlate[Sbr_IN_dCapIndex].tData.dTotalCaps > 1) AND (TMP_dNextCap > 0) THEN
   	JSR(sbrCheckConvoyZCDestination,5,TMP_dNextCap,Sbr_INO_DestinationLite,Sbr_IN_DestinationCullet,Sbr_INO_xAtLeastOneForDestination,Sbr_INO_xAtLeastOneToCullet,Sbr_INO_xAtLeastOneForDestination,Sbr_INO_xAllLiteToCullet);
   END_IF;
   
   RET(Sbr_INO_xALLForDestination,Sbr_INO_xAtLeastOneToCullet);
   
END_ROUTINE

ROUTINE sbrConvDataLineToSL   (* structured text *)
   
   //Input
   SBR(Sbr_INO_tConvoyCap_ZC,Sbr_INO_tConvoy_SL,Sbr_IN_dCapIndex);